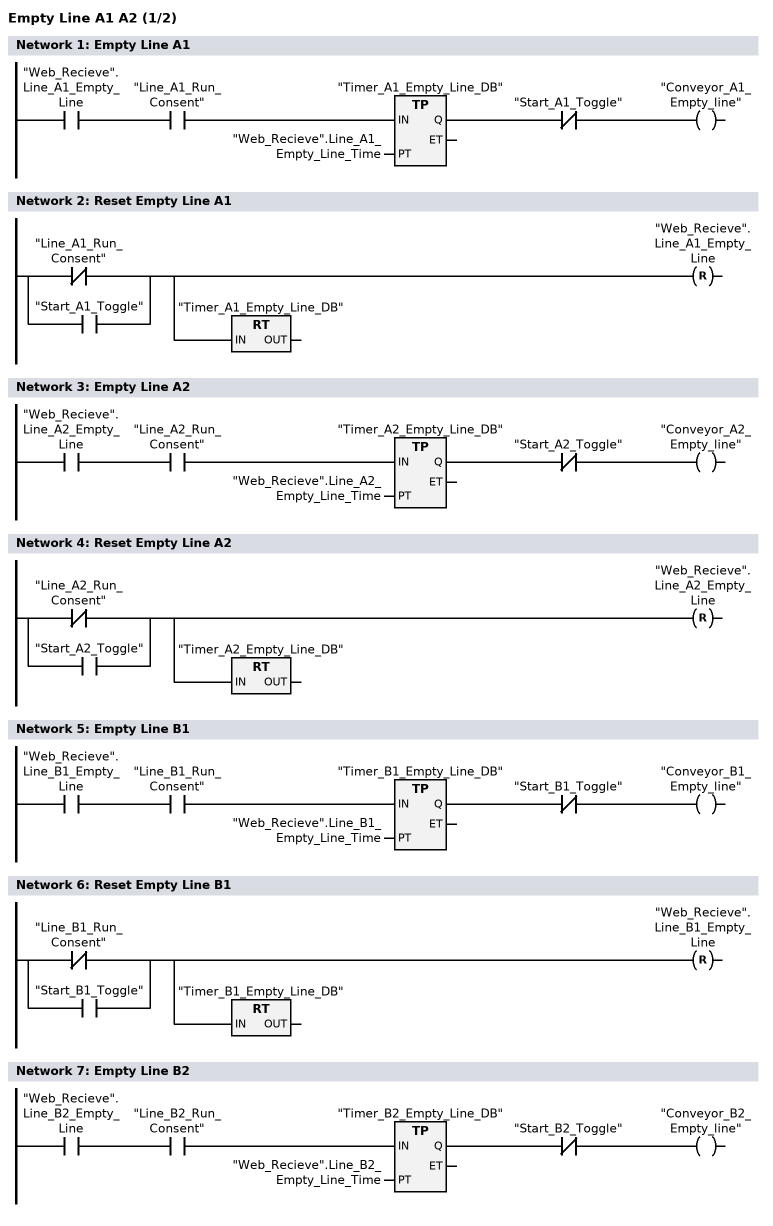
   "Timer_A1_Empty_Line_DB".TP(IN := "Web_Recieve".Line_A1_Empty_Line AND "Line_A1_Run_Consent",
                           PT := "Web_Recieve".Line_A1_Empty_Line_Time);
   "Conveyor_A1_Empty_line" := "Timer_A1_Empty_Line_DB".Q AND NOT "Start_A1_Toggle";
END_REGION

REGION Network 2: Reset Empty Line A1
   RUNG wire#powerrail
      I_Contact( "Line_A1_Run_Consent" )
      wire#w1
      R_Coil( "Web_Recieve".Line_A1_Empty_Line )
   END_RUNG
   RUNG wire#powerrail
      Contact( "Start_A1_Toggle" )
   END_RUNG wire#w1
   RUNG wire#w1
      RT_Coil( "Timer_A1_Empty_Line_DB" )
   END_RUNG
   // the same network as SCL:
   #_w1 := NOT "Line_A1_Run_Consent" OR "Start_A1_Toggle";
   IF #_w1 THEN
       "Web_Recieve".Line_A1_Empty_Line := FALSE;
       RESET_TIMER("Timer_A1_Empty_Line_DB");
   END_IF;
END_REGION

REGION Network 3: Empty Line A2
   "Timer_A2_Empty_Line_DB".TP(IN := "Web_Recieve".Line_A2_Empty_Line AND "Line_A2_Run_Consent",
                           PT := "Web_Recieve".Line_A2_Empty_Line_Time);
   "Conveyor_A2_Empty_line" := "Timer_A2_Empty_Line_DB".Q AND NOT "Start_A2_Toggle";
END_REGION

REGION Network 4: Reset Empty Line A2
   RUNG wire#powerrail
      I_Contact( "Line_A2_Run_Consent" )
      wire#w1
      R_Coil( "Web_Recieve".Line_A2_Empty_Line )
   END_RUNG
   RUNG wire#powerrail
      Contact( "Start_A2_Toggle" )
   END_RUNG wire#w1
   RUNG wire#w1
      RT_Coil( "Timer_A2_Empty_Line_DB" )
   END_RUNG
   // the same network as SCL:
   #_w1 := NOT "Line_A2_Run_Consent" OR "Start_A2_Toggle";
   IF #_w1 THEN
       "Web_Recieve".Line_A2_Empty_Line := FALSE;
       RESET_TIMER("Timer_A2_Empty_Line_DB");
   END_IF;
END_REGION

REGION Network 5: Empty Line B1
   "Timer_B1_Empty_Line_DB".TP(IN := "Web_Recieve".Line_B1_Empty_Line AND "Line_B1_Run_Consent",
                           PT := "Web_Recieve".Line_B1_Empty_Line_Time);
   "Conveyor_B1_Empty_line" := "Timer_B1_Empty_Line_DB".Q AND NOT "Start_B1_Toggle";
END_REGION

REGION Network 6: Reset Empty Line B1
   RUNG wire#powerrail
      I_Contact( "Line_B1_Run_Consent" )
      wire#w1
      R_Coil( "Web_Recieve".Line_B1_Empty_Line )
   END_RUNG
   RUNG wire#powerrail
      Contact( "Start_B1_Toggle" )
   END_RUNG wire#w1
   RUNG wire#w1
      RT_Coil( "Timer_B1_Empty_Line_DB" )
   END_RUNG
   // the same network as SCL:
   #_w1 := NOT "Line_B1_Run_Consent" OR "Start_B1_Toggle";
   IF #_w1 THEN
       "Web_Recieve".Line_B1_Empty_Line := FALSE;
       RESET_TIMER("Timer_B1_Empty_Line_DB");
   END_IF;
END_REGION

REGION Network 7: Empty Line B2
   "Timer_B2_Empty_Line_DB".TP(IN := "Web_Recieve".Line_B2_Empty_Line AND "Line_B2_Run_Consent",
                           PT := "Web_Recieve".Line_B2_Empty_Line_Time);
   "Conveyor_B2_Empty_line" := "Timer_B2_Empty_Line_DB".Q AND NOT "Start_B2_Toggle";
END_REGION

REGION Network 8: Reset Empty Line B2
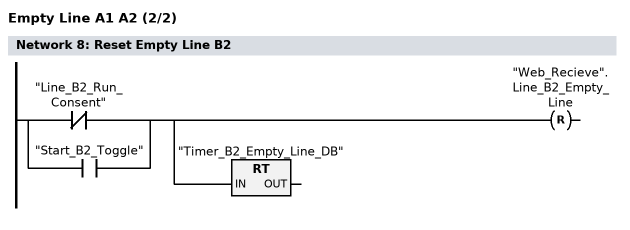
   RUNG wire#powerrail
      I_Contact( "Line_B2_Run_Consent" )
      wire#w1
      R_Coil( "Web_Recieve".Line_B2_Empty_Line )
   END_RUNG
   RUNG wire#powerrail
      Contact( "Start_B2_Toggle" )
   END_RUNG wire#w1
   RUNG wire#w1
      RT_Coil( "Timer_B2_Empty_Line_DB" )
   END_RUNG
   // the same network as SCL:
   #_w1 := NOT "Line_B2_Run_Consent" OR "Start_B2_Toggle";
   IF #_w1 THEN
       "Web_Recieve".Line_B2_Empty_Line := FALSE;
       RESET_TIMER("Timer_B2_Empty_Line_DB");
   END_IF;
END_REGION
END_FUNCTION_BLOCK

FUNCTION_BLOCK "Empty Line B1 B2"   // FB14, LAD
{ S7_Optimized_Access := 'TRUE' }
VERSION : 0.1
BEGIN

REGION Network 1
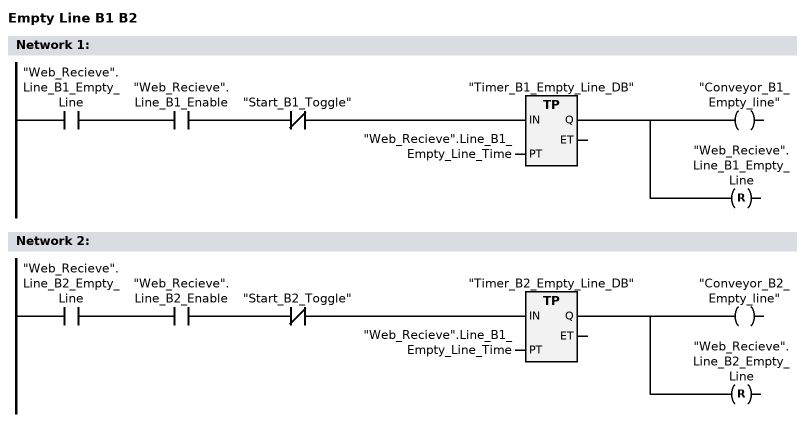
   "Timer_B1_Empty_Line_DB".TP(IN := "Web_Recieve".Line_B1_Empty_Line AND "Web_Recieve".Line_B1_Enable AND NOT "Start_B1_Toggle",
                           PT := "Web_Recieve".Line_B1_Empty_Line_Time);
   "Conveyor_B1_Empty_line" := "Timer_B1_Empty_Line_DB".Q;
   IF "Timer_B1_Empty_Line_DB".Q THEN "Web_Recieve".Line_B1_Empty_Line := FALSE; END_IF;
END_REGION

REGION Network 2
   "Timer_B2_Empty_Line_DB".TP(IN := "Web_Recieve".Line_B2_Empty_Line AND "Web_Recieve".Line_B2_Enable AND NOT "Start_B2_Toggle",
                           PT := "Web_Recieve".Line_B1_Empty_Line_Time);
   "Conveyor_B2_Empty_line" := "Timer_B2_Empty_Line_DB".Q;
   IF "Timer_B2_Empty_Line_DB".Q THEN "Web_Recieve".Line_B2_Empty_Line := FALSE; END_IF;
END_REGION
END_FUNCTION_BLOCK

FUNCTION_BLOCK "SaveDataToDataBlock A1"   // FB15, LAD
{ S7_Optimized_Access := 'TRUE' }
VERSION : 0.1
   VAR_TEMP
      Busytemp : Bool;
      returnValueTemp : DInt;
   END_VAR
BEGIN

REGION Network 1: Line_A1_Conveyer_on_Time Save
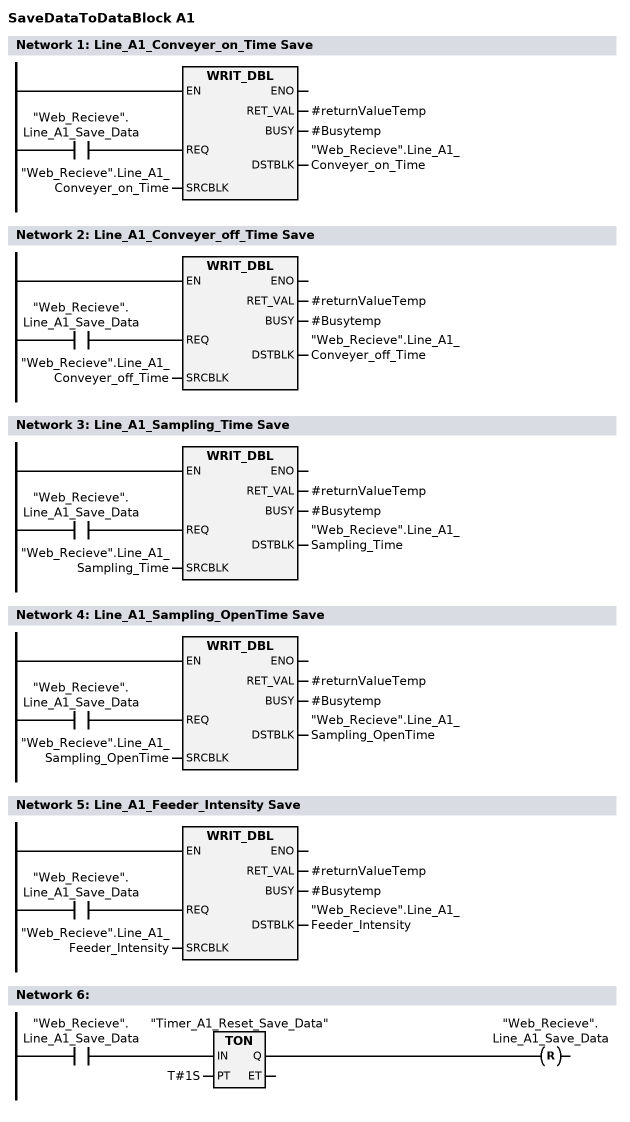
   #returnValueTemp := WRIT_DBL(REQ := "Web_Recieve".Line_A1_Save_Data,
                           SRCBLK := "Web_Recieve".Line_A1_Conveyer_on_Time,
                           BUSY => #Busytemp,
                           DSTBLK => "Web_Recieve".Line_A1_Conveyer_on_Time);
END_REGION

REGION Network 2: Line_A1_Conveyer_off_Time Save
   #returnValueTemp := WRIT_DBL(REQ := "Web_Recieve".Line_A1_Save_Data,
                           SRCBLK := "Web_Recieve".Line_A1_Conveyer_off_Time,
                           BUSY => #Busytemp,
                           DSTBLK => "Web_Recieve".Line_A1_Conveyer_off_Time);
END_REGION

REGION Network 3: Line_A1_Sampling_Time Save
   #returnValueTemp := WRIT_DBL(REQ := "Web_Recieve".Line_A1_Save_Data,
                           SRCBLK := "Web_Recieve".Line_A1_Sampling_Time,
                           BUSY => #Busytemp,
                           DSTBLK => "Web_Recieve".Line_A1_Sampling_Time);
END_REGION

REGION Network 4: Line_A1_Sampling_OpenTime Save
   #returnValueTemp := WRIT_DBL(REQ := "Web_Recieve".Line_A1_Save_Data,
                           SRCBLK := "Web_Recieve".Line_A1_Sampling_OpenTime,
                           BUSY => #Busytemp,
                           DSTBLK => "Web_Recieve".Line_A1_Sampling_OpenTime);
END_REGION

REGION Network 5: Line_A1_Feeder_Intensity Save
   #returnValueTemp := WRIT_DBL(REQ := "Web_Recieve".Line_A1_Save_Data,
                           SRCBLK := "Web_Recieve".Line_A1_Feeder_Intensity,
                           BUSY => #Busytemp,
                           DSTBLK => "Web_Recieve".Line_A1_Feeder_Intensity);
END_REGION

REGION Network 6
   "Timer_A1_Reset_Save_Data".TON(IN := "Web_Recieve".Line_A1_Save_Data, PT := T#1S);
   IF "Timer_A1_Reset_Save_Data".Q THEN "Web_Recieve".Line_A1_Save_Data := FALSE; END_IF;
END_REGION
END_FUNCTION_BLOCK

FUNCTION_BLOCK "SaveDataToDataBlock A2"   // FB16, LAD
{ S7_Optimized_Access := 'TRUE' }
VERSION : 0.1
   VAR_TEMP
      Busytemp : Bool;
      returnValueTemp : DInt;
   END_VAR
BEGIN

REGION Network 1: Line_A2_Conveyer_on_Time Save
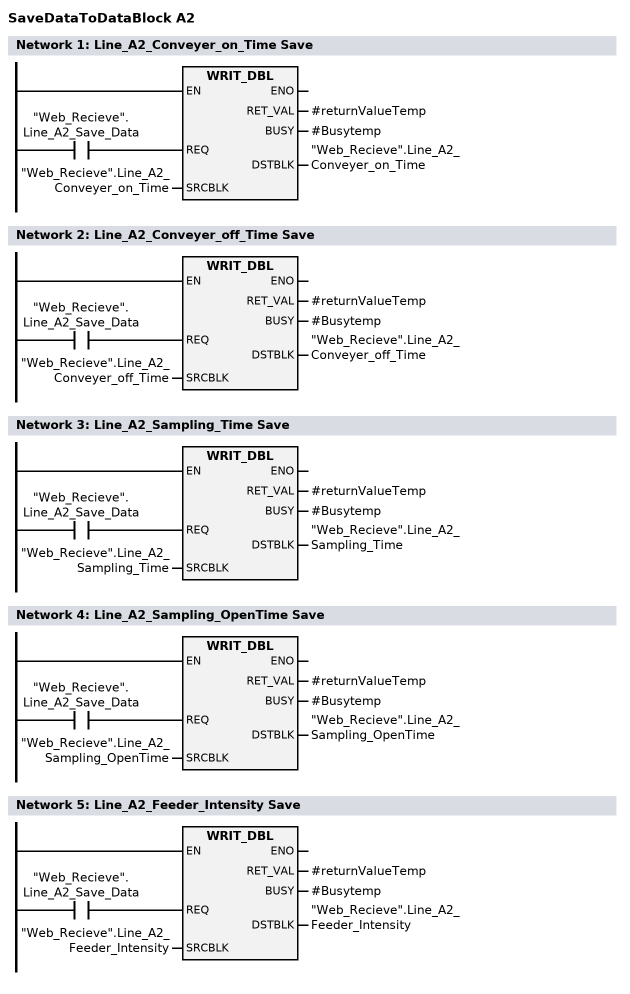
   #returnValueTemp := WRIT_DBL(REQ := "Web_Recieve".Line_A2_Save_Data,
                           SRCBLK := "Web_Recieve".Line_A2_Conveyer_on_Time,
                           BUSY => #Busytemp,
                           DSTBLK => "Web_Recieve".Line_A2_Conveyer_on_Time);
END_REGION

REGION Network 2: Line_A2_Conveyer_off_Time Save
   #returnValueTemp := WRIT_DBL(REQ := "Web_Recieve".Line_A2_Save_Data,
                           SRCBLK := "Web_Recieve".Line_A2_Conveyer_off_Time,
                           BUSY => #Busytemp,
                           DSTBLK => "Web_Recieve".Line_A2_Conveyer_off_Time);
END_REGION

REGION Network 3: Line_A2_Sampling_Time Save
   #returnValueTemp := WRIT_DBL(REQ := "Web_Recieve".Line_A2_Save_Data,
                           SRCBLK := "Web_Recieve".Line_A2_Sampling_Time,
                           BUSY => #Busytemp,
                           DSTBLK => "Web_Recieve".Line_A2_Sampling_Time);
END_REGION

REGION Network 4: Line_A2_Sampling_OpenTime Save
   #returnValueTemp := WRIT_DBL(REQ := "Web_Recieve".Line_A2_Save_Data,
                           SRCBLK := "Web_Recieve".Line_A2_Sampling_OpenTime,
                           BUSY => #Busytemp,
                           DSTBLK => "Web_Recieve".Line_A2_Sampling_OpenTime);
END_REGION

REGION Network 5: Line_A2_Feeder_Intensity Save
   #returnValueTemp := WRIT_DBL(REQ := "Web_Recieve".Line_A2_Save_Data,
                           SRCBLK := "Web_Recieve".Line_A2_Feeder_Intensity,
                           BUSY => #Busytemp,
                           DSTBLK => "Web_Recieve".Line_A2_Feeder_Intensity);
END_REGION
END_FUNCTION_BLOCK

FUNCTION_BLOCK "SaveDataToDataBlock B2"   // FB17, LAD
{ S7_Optimized_Access := 'TRUE' }
VERSION : 0.1
   VAR_TEMP
      Busytemp : Bool;
      returnValueTemp : DInt;
   END_VAR
BEGIN

REGION Network 1: Line_B2_Conveyer_on_Time Save
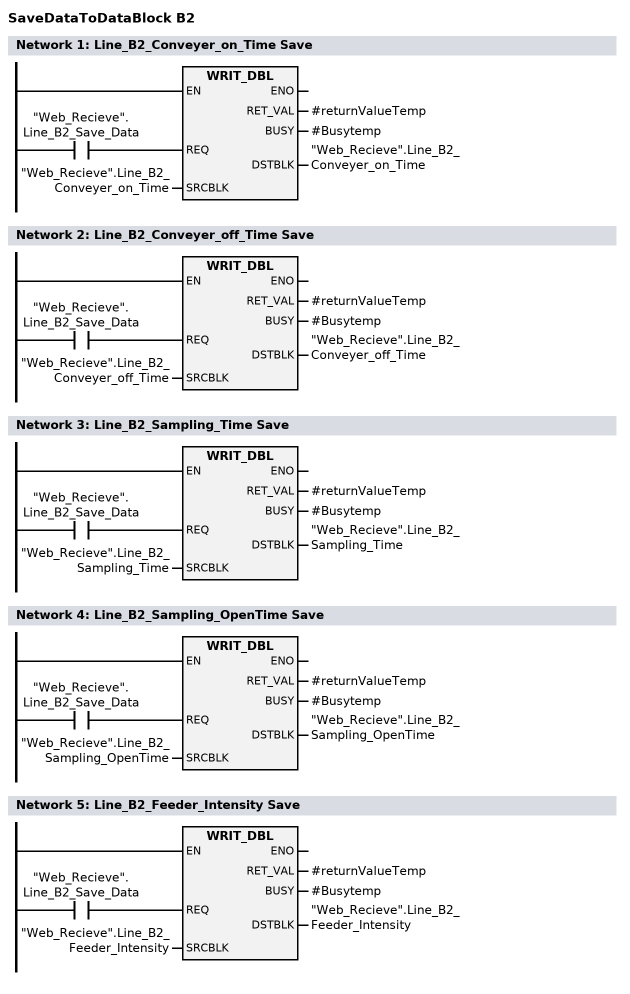
   #returnValueTemp := WRIT_DBL(REQ := "Web_Recieve".Line_B2_Save_Data,
                           SRCBLK := "Web_Recieve".Line_B2_Conveyer_on_Time,
                           BUSY => #Busytemp,
                           DSTBLK => "Web_Recieve".Line_B2_Conveyer_on_Time);
END_REGION

REGION Network 2: Line_B2_Conveyer_off_Time Save
   #returnValueTemp := WRIT_DBL(REQ := "Web_Recieve".Line_B2_Save_Data,
                           SRCBLK := "Web_Recieve".Line_B2_Conveyer_off_Time,
                           BUSY => #Busytemp,
                           DSTBLK => "Web_Recieve".Line_B2_Conveyer_off_Time);
END_REGION

REGION Network 3: Line_B2_Sampling_Time Save
   #returnValueTemp := WRIT_DBL(REQ := "Web_Recieve".Line_B2_Save_Data,
                           SRCBLK := "Web_Recieve".Line_B2_Sampling_Time,
                           BUSY => #Busytemp,
                           DSTBLK => "Web_Recieve".Line_B2_Sampling_Time);
END_REGION

REGION Network 4: Line_B2_Sampling_OpenTime Save
   #returnValueTemp := WRIT_DBL(REQ := "Web_Recieve".Line_B2_Save_Data,
                           SRCBLK := "Web_Recieve".Line_B2_Sampling_OpenTime,
                           BUSY => #Busytemp,
                           DSTBLK => "Web_Recieve".Line_B2_Sampling_OpenTime);
END_REGION

REGION Network 5: Line_B2_Feeder_Intensity Save
   #returnValueTemp := WRIT_DBL(REQ := "Web_Recieve".Line_B2_Save_Data,
                           SRCBLK := "Web_Recieve".Line_B2_Feeder_Intensity,
                           BUSY => #Busytemp,
                           DSTBLK => "Web_Recieve".Line_B2_Feeder_Intensity);
END_REGION
END_FUNCTION_BLOCK

FUNCTION_BLOCK "SaveDataToDataBlock B1"   // FB18, LAD
{ S7_Optimized_Access := 'TRUE' }
VERSION : 0.1
   VAR_TEMP
      Busytemp : Bool;
      returnValueTemp : DInt;
   END_VAR
BEGIN

REGION Network 1: Line_B1_Conveyer_on_Time Save
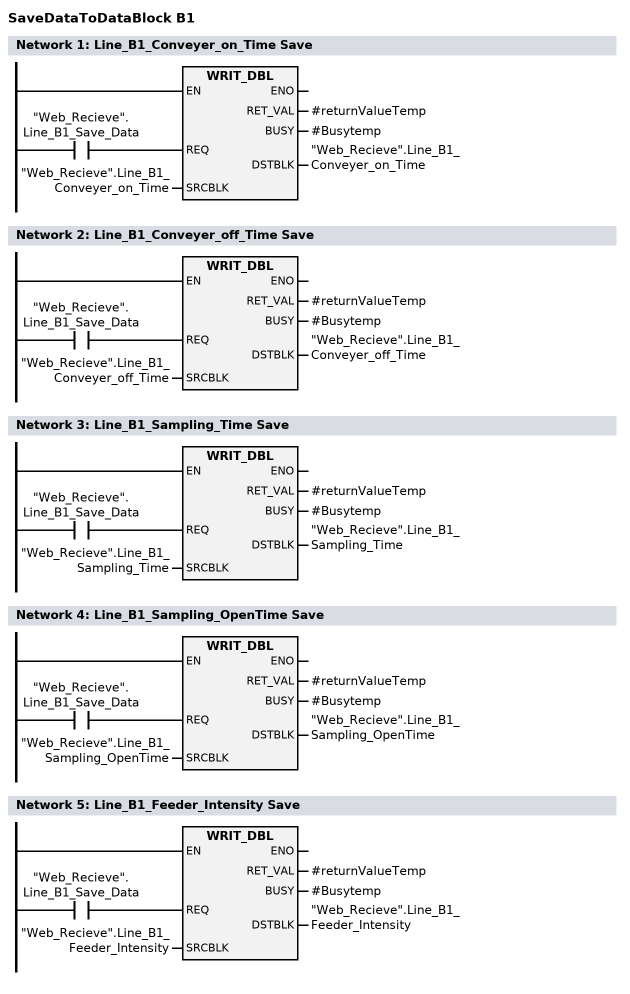
   #returnValueTemp := WRIT_DBL(REQ := "Web_Recieve".Line_B1_Save_Data,
                           SRCBLK := "Web_Recieve".Line_B1_Conveyer_on_Time,
                           BUSY => #Busytemp,
                           DSTBLK => "Web_Recieve".Line_B1_Conveyer_on_Time);
END_REGION

REGION Network 2: Line_B1_Conveyer_off_Time Save
   #returnValueTemp := WRIT_DBL(REQ := "Web_Recieve".Line_B1_Save_Data,
                           SRCBLK := "Web_Recieve".Line_B1_Conveyer_off_Time,
                           BUSY => #Busytemp,
                           DSTBLK => "Web_Recieve".Line_B1_Conveyer_off_Time);
END_REGION

REGION Network 3: Line_B1_Sampling_Time Save
   #returnValueTemp := WRIT_DBL(REQ := "Web_Recieve".Line_B1_Save_Data,
                           SRCBLK := "Web_Recieve".Line_B1_Sampling_Time,
                           BUSY => #Busytemp,
                           DSTBLK => "Web_Recieve".Line_B1_Sampling_Time);
END_REGION

REGION Network 4: Line_B1_Sampling_OpenTime Save
   #returnValueTemp := WRIT_DBL(REQ := "Web_Recieve".Line_B1_Save_Data,
                           SRCBLK := "Web_Recieve".Line_B1_Sampling_OpenTime,
                           BUSY => #Busytemp,
                           DSTBLK => "Web_Recieve".Line_B1_Sampling_OpenTime);
END_REGION

REGION Network 5: Line_B1_Feeder_Intensity Save
   #returnValueTemp := WRIT_DBL(REQ := "Web_Recieve".Line_B1_Save_Data,
                           SRCBLK := "Web_Recieve".Line_B1_Feeder_Intensity,
                           BUSY => #Busytemp,
                           DSTBLK => "Web_Recieve".Line_B1_Feeder_Intensity);
END_REGION
END_FUNCTION_BLOCK

ORGANIZATION_BLOCK "Main"   // OB1, LAD, ProgramCycle
TITLE = "Main Program Sweep (Cycle)"
{ S7_Optimized_Access := 'TRUE' }
VERSION : 0.1
   VAR_INPUT
      Initial_Call : Bool;   // Initial call of this OB
      Remanence : Bool;   // =True, if remanent data are available
   END_VAR
   VAR_TEMP
      TEMP : Int;
      clkRetVal : Int;
      newt : Int;
      ModbusDone : Bool;
      ModbusError : Bool;
      ModbusStatus : Word;
      ModbusWriteDone : Bool;
   END_VAR
BEGIN

REGION Network 1: Web data WWW
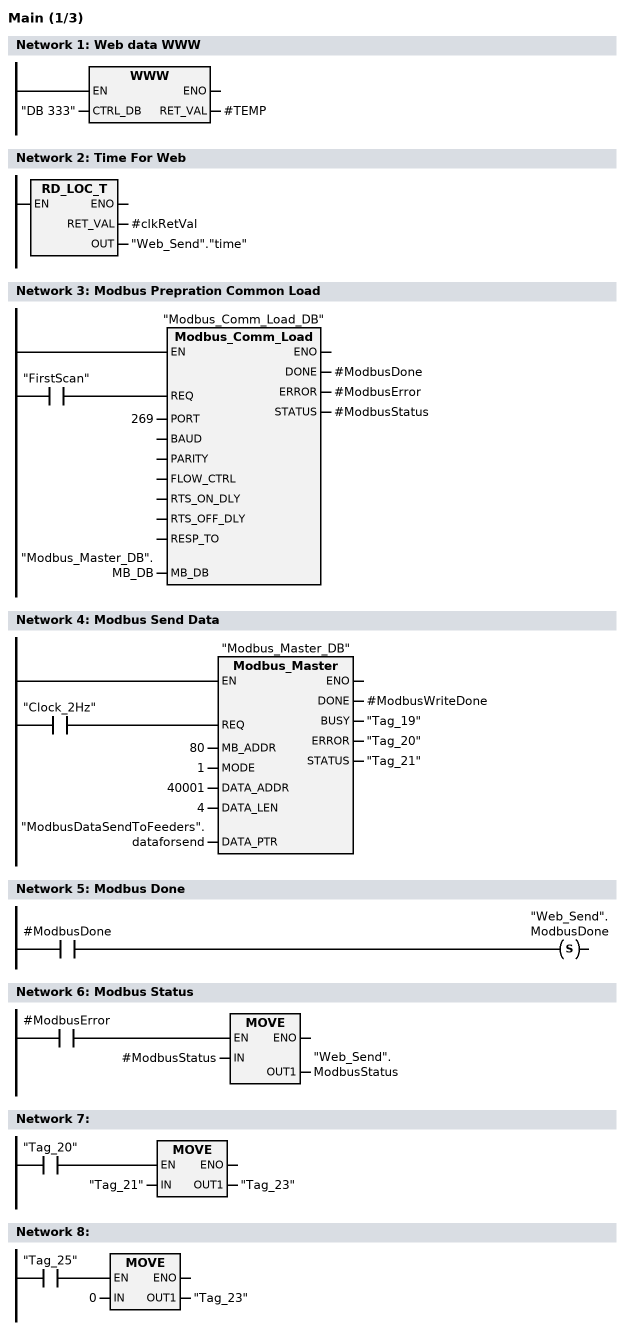
   #TEMP := WWW(CTRL_DB := "DB 333");
END_REGION

REGION Network 2: Time For Web
   #clkRetVal := RD_LOC_T(OUT => "Web_Send"."time");
END_REGION

REGION Network 3: Modbus Prepration Common Load
   "Modbus_Comm_Load_DB"(REQ := "FirstScan",   // Modbus_Comm_Load
                         PORT := 269,
                         MB_DB := "Modbus_Master_DB".MB_DB,
                         DONE => #ModbusDone,
                         ERROR => #ModbusError,
                         STATUS => #ModbusStatus);
END_REGION

REGION Network 4: Modbus Send Data
   "Modbus_Master_DB"(REQ := "Clock_2Hz",   // Modbus_Master
                      MB_ADDR := 80,
                      MODE := 1,
                      DATA_ADDR := 40001,
                      DATA_LEN := 4,
                      DATA_PTR := "ModbusDataSendToFeeders".dataforsend,
                      DONE => #ModbusWriteDone,
                      BUSY => "Tag_19",
                      ERROR => "Tag_20",
                      STATUS => "Tag_21");
END_REGION

REGION Network 5: Modbus Done
   RUNG wire#powerrail
      Contact( #ModbusDone )
      S_Coil( "Web_Send".ModbusDone )
   END_RUNG
   // the same network as SCL:
   IF #ModbusDone THEN "Web_Send".ModbusDone := TRUE; END_IF;
END_REGION

REGION Network 6: Modbus Status
   RUNG wire#powerrail
      Contact( #ModbusError )
      Move(in := #ModbusStatus, out1 => "Web_Send".ModbusStatus)
   END_RUNG
   // the same network as SCL:
   IF #ModbusError THEN "Web_Send".ModbusStatus := #ModbusStatus; END_IF;
END_REGION

REGION Network 7
   RUNG wire#powerrail
      Contact( "Tag_20" )
      Move(in := "Tag_21", out1 => "Tag_23")
   END_RUNG
   // the same network as SCL:
   IF "Tag_20" THEN "Tag_23" := "Tag_21"; END_IF;
END_REGION

REGION Network 8
   RUNG wire#powerrail
      Contact( "Tag_25" )
      Move(in := 0, out1 => "Tag_23")
   END_RUNG
   // the same network as SCL:
   IF "Tag_25" THEN "Tag_23" := 0; END_IF;
END_REGION

REGION Network 9
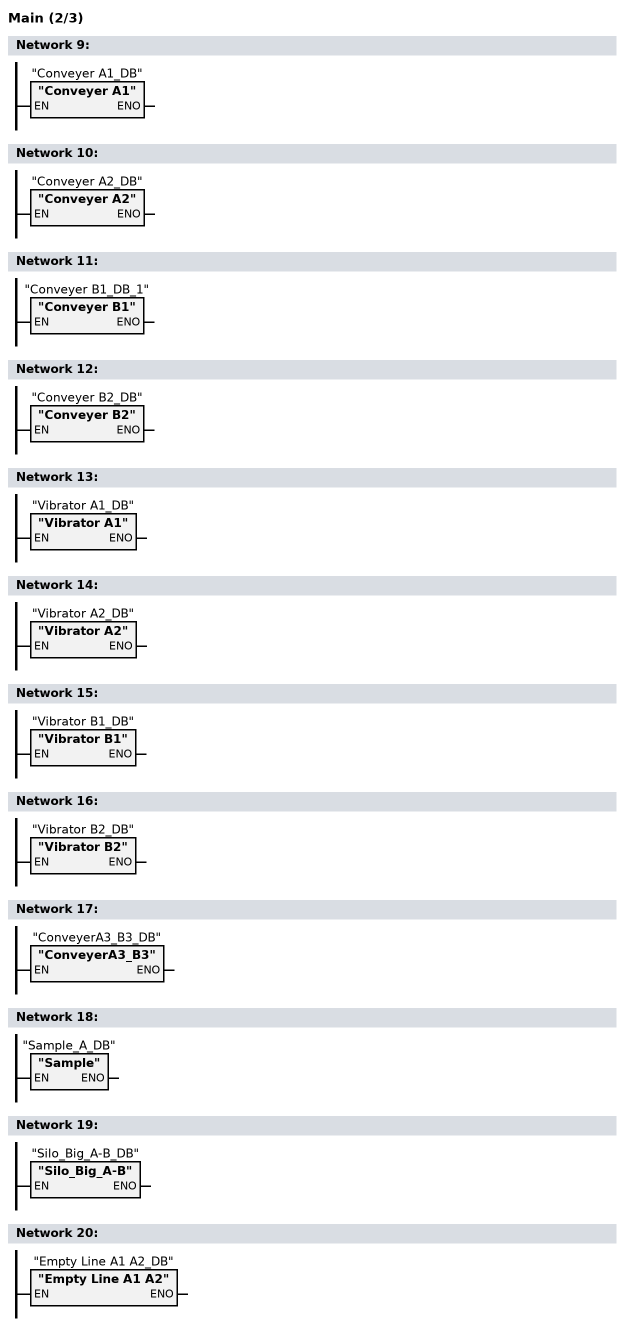
   RUNG wire#powerrail
      "Conveyer A1_DB"()
   END_RUNG
   // the same network as SCL:
   "Conveyer A1_DB"();   // "Conveyer A1"
END_REGION

REGION Network 10
   RUNG wire#powerrail
      "Conveyer A2_DB"()
   END_RUNG
   // the same network as SCL:
   "Conveyer A2_DB"();   // "Conveyer A2"
END_REGION

REGION Network 11
   RUNG wire#powerrail
      "Conveyer B1_DB_1"()
   END_RUNG
   // the same network as SCL:
   "Conveyer B1_DB_1"();   // "Conveyer B1"
END_REGION

REGION Network 12
   RUNG wire#powerrail
      "Conveyer B2_DB"()
   END_RUNG
   // the same network as SCL:
   "Conveyer B2_DB"();   // "Conveyer B2"
END_REGION

REGION Network 13
   RUNG wire#powerrail
      "Vibrator A1_DB"()
   END_RUNG
   // the same network as SCL:
   "Vibrator A1_DB"();   // "Vibrator A1"
END_REGION

REGION Network 14
   RUNG wire#powerrail
      "Vibrator A2_DB"()
   END_RUNG
   // the same network as SCL:
   "Vibrator A2_DB"();   // "Vibrator A2"
END_REGION

REGION Network 15
   RUNG wire#powerrail
      "Vibrator B1_DB"()
   END_RUNG
   // the same network as SCL:
   "Vibrator B1_DB"();   // "Vibrator B1"
END_REGION

REGION Network 16
   RUNG wire#powerrail
      "Vibrator B2_DB"()
   END_RUNG
   // the same network as SCL:
   "Vibrator B2_DB"();   // "Vibrator B2"
END_REGION

REGION Network 17
   RUNG wire#powerrail
      "ConveyerA3_B3_DB"()
   END_RUNG
   // the same network as SCL:
   "ConveyerA3_B3_DB"();   // "ConveyerA3_B3"
END_REGION

REGION Network 18
   RUNG wire#powerrail
      "Sample_A_DB"()
   END_RUNG
   // the same network as SCL:
   "Sample_A_DB"();   // "Sample"
END_REGION

REGION Network 19
   RUNG wire#powerrail
      "Silo_Big_A-B_DB"()
   END_RUNG
   // the same network as SCL:
   "Silo_Big_A-B_DB"();   // "Silo_Big_A-B"
END_REGION

REGION Network 20
   RUNG wire#powerrail
      "Empty Line A1 A2_DB"()
   END_RUNG
   // the same network as SCL:
   "Empty Line A1 A2_DB"();   // "Empty Line A1 A2"
END_REGION

REGION Network 21
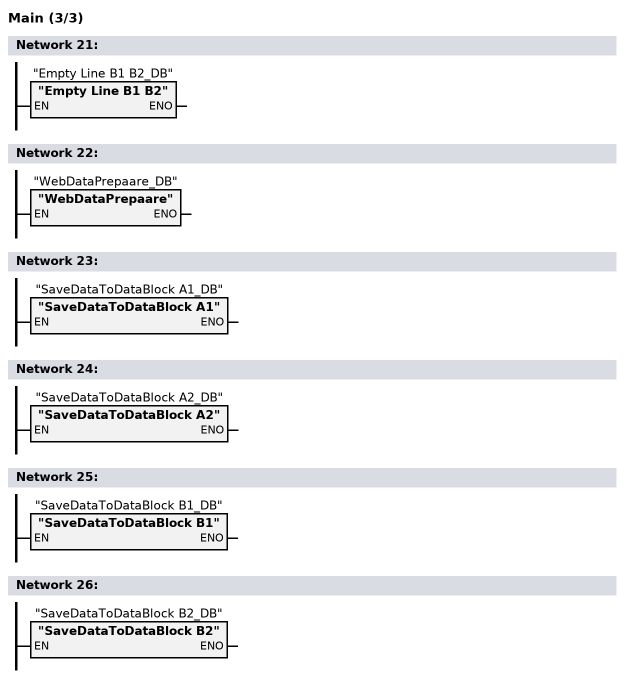
   RUNG wire#powerrail
      "Empty Line B1 B2_DB"()
   END_RUNG
   // the same network as SCL:
   "Empty Line B1 B2_DB"();   // "Empty Line B1 B2"
END_REGION

REGION Network 22
   RUNG wire#powerrail
      "WebDataPrepaare_DB"()
   END_RUNG
   // the same network as SCL:
   "WebDataPrepaare_DB"();   // "WebDataPrepaare"
END_REGION

REGION Network 23
   RUNG wire#powerrail
      "SaveDataToDataBlock A1_DB"()
   END_RUNG
   // the same network as SCL:
   "SaveDataToDataBlock A1_DB"();   // "SaveDataToDataBlock A1"
END_REGION

REGION Network 24
   RUNG wire#powerrail
      "SaveDataToDataBlock A2_DB"()
   END_RUNG
   // the same network as SCL:
   "SaveDataToDataBlock A2_DB"();   // "SaveDataToDataBlock A2"
END_REGION

REGION Network 25
   RUNG wire#powerrail
      "SaveDataToDataBlock B1_DB"()
   END_RUNG
   // the same network as SCL:
   "SaveDataToDataBlock B1_DB"();   // "SaveDataToDataBlock B1"
END_REGION

REGION Network 26
   RUNG wire#powerrail
      "SaveDataToDataBlock B2_DB"()
   END_RUNG
   // the same network as SCL:
   "SaveDataToDataBlock B2_DB"();   // "SaveDataToDataBlock B2"
END_REGION
END_ORGANIZATION_BLOCK